// TIA Portal project "Tes simulation extract_V15.1" (V15.1)

(* hardware
DEVICE "S71500/ET200MP station_1"  S7-1500 station
   slot 0: "Rail_0"  Rack  6ES7 590-1***0-0AA0
   slot 1: "PLC_1"  CPU 1511-1 PN  6ES7 511-1AK01-0AB0  V2.1
      slot 3: "CPU display_1"  6ES7591-1AA00-0AA0
DEVICE "PC station"  SIMATIC PC station
   slot 0: "PC station"  Rail  SIMATIC PC-Station  V1.0
      slot 125: "Stationmanager"  Station_Manager  V6.0.4
   slot 1: "IE general_1"  IE General  IE_CP  V8.2.0
   slot 2: "HMI_RT_1"  WinCC RT Advanced  6AV2 104-0xxxx-xxxx  15.1.0.0
      slot 33792: "Host interface"  Host interface
*)

// ===== PLC "PLC_1"  CPU 1511-1 PN =====

VAR_GLOBAL   // PLC tag table "Default tag table"
   "Clock_Byte" AT %MB0 : Byte;
   "Clock_10Hz" AT %M0.0 : Bool;
   "Clock_5Hz" AT %M0.1 : Bool;
   "Clock_2.5Hz" AT %M0.2 : Bool;
   "Clock_2Hz" AT %M0.3 : Bool;
   "Clock_1.25Hz" AT %M0.4 : Bool;
   "Clock_1Hz" AT %M0.5 : Bool;
   "Clock_0.625Hz" AT %M0.6 : Bool;
   "Clock_0.5Hz" AT %M0.7 : Bool;
   "Start Preparation V1" AT %M100.0 : Bool;
   "Pressure Vesel" AT %MW200 : Word;
   "Pressure Steam" AT %MW230 : Int;
   "Tag_3" AT %MW1 : Word;
   "Tag_4" AT %MB1 : Byte;
   "Tag_5" AT %T1 : Timer;
   "Tag_2" AT %T2 : Timer;
   "Tag_6" AT %MB26 : Byte;
   "Tag_7" AT %T3 : Timer;
   "Tag_8" AT %T4 : Timer;
   "Tag_9" AT %T5 : Timer;
   "Tag_10" AT %M100.1 : Bool;
   "Tag_11" AT %T6 : Timer;
   "Tag_12" AT %T7 : Timer;
   "START Proses" AT %M100.2 : Bool;
   "Tag_13" AT %T8 : Timer;
   "Tag_14" AT %MB4 : Byte;
   "Tag_15" AT %T9 : Timer;
   "Tag_16" AT %MB8 : Byte;
   "Tag_17" AT %MB6 : Byte;
   "Tag_18" AT %T10 : Timer;
   "START SUPPLY" AT %M100.3 : Bool;
   "Tag_20" AT %T11 : Timer;
   "TEMP SENSOR 1" AT %MW164 : Word;
   "Tag_21" AT %T12 : Timer;
   "TEMP SENSOR 2" AT %MW166 : Int;
   "Tag_22" AT %MB30 : Byte;
   "START PROSES V1" AT %M100.4 : Bool;
   "Tag_19" AT %MW2 : Int;
   "TEMPERATURE VESSEL 1" AT %MW240 : Int;
   "Tag_23" AT %MB2 : Byte;
   "Tag_24" AT %T13 : Timer;
   "Tag_25" AT %T14 : Timer;
   "Tag_26" AT %T15 : Timer;
   "Tag_27" AT %T16 : Timer;
   "Tag_28" AT %T17 : Timer;
   "Tag_29" AT %T18 : Timer;
   "Tag_30" AT %T19 : Timer;
   "Tag_31" AT %T20 : Timer;
   "Tag_32" AT %T21 : Timer;
   "Tag_33" AT %T22 : Timer;
   "Count Preparation V1" AT %MW120 : Int;
   "Count Step Proses V1" AT %MW140 : Int;
   "START TRANSFER" AT %M100.5 : Bool;
   "Tag_36" AT %M30.4 : Bool;
   "Tag_37" AT %T23 : Timer;
   "Tag_38" AT %T24 : Timer;
   "Tag_39" AT %T35 : Timer;
   "Tag_40" AT %T25 : Timer;
   "Tag_41" AT %T26 : Timer;
   "START PROSES V2" AT %M100.6 : Bool;
   "Pressure Vessel 2" AT %MW202 : Int;
   "TEMPERATURE VESSEL 2" AT %MW242 : Int;
   "Tag_42" AT %T27 : Timer;
   "Tag_43" AT %T28 : Timer;
   "Tag_44" AT %T29 : Timer;
   "Tag_45" AT %T30 : Timer;
   "Tag_46" AT %T31 : Timer;
   "Tag_47" AT %T32 : Timer;
   "Tag_48" AT %T33 : Timer;
   "Tag_49" AT %T34 : Timer;
   "Tag_50" AT %T36 : Timer;
   "Count Step Proses V2" AT %MW142 : Int;
   "Tag_52" AT %MB5 : Byte;
   "Start Preparation V7" AT %M102.0 : Bool;
   "Tag_54" AT %M102.1 : Bool;
   "START PROSES V3" AT %M100.7 : Bool;
   "Tag_55" AT %T38 : Timer;
   "Pressure Vessel 3" AT %MW204 : Int;
   "TEMPERATURE VESSEL 3" AT %MW244 : Int;
   "Tag_56" AT %T39 : Timer;
   "Tag_57" AT %T40 : Timer;
   "Tag_58" AT %T41 : Timer;
   "Tag_59" AT %T42 : Timer;
   "Tag_60" AT %T43 : Timer;
   "Tag_61" AT %T44 : Timer;
   "Tag_62" AT %T45 : Timer;
   "Tag_63" AT %T46 : Timer;
   "Tag_64" AT %T47 : Timer;
   "Count Step Proses V3" AT %MW144 : Int;
   "Tag_66" AT %MB9 : Byte;
   "Tag_67" AT %M102.2 : Bool;
   "Start Proses V4" AT %M101.0 : Bool;
   "Pressure Vessel 4" AT %MW206 : Int;
   "Tag_69" AT %T48 : Timer;
   "TEMPERATURE VESSEL 4" AT %MW246 : Int;
   "Tag_70" AT %T49 : Timer;
   "Tag_71" AT %T50 : Timer;
   "Tag_72" AT %T51 : Timer;
   "Tag_73" AT %T52 : Timer;
   "Tag_74" AT %T53 : Timer;
   "Tag_75" AT %T54 : Timer;
   "Tag_76" AT %T55 : Timer;
   "Tag_77" AT %T56 : Timer;
   "Tag_78" AT %T57 : Timer;
   "Count Step Proses V4" AT %MW146 : Int;
   "Tag_80" AT %MB12 : Byte;
   "Tag_81" AT %MB13 : Byte;
   "Pressure vessel 5" AT %MW208 : Int;
   "TEMPERATURE VESSEL 5" AT %MW248 : Int;
   "START PROSES V5" AT %M101.1 : Bool;
   "Tag_82" AT %M102.3 : Bool;
   "Tag_83" AT %T58 : Timer;
   "Tag_84" AT %T59 : Timer;
   "Tag_85" AT %T60 : Timer;
   "Tag_86" AT %T61 : Timer;
   "Tag_87" AT %T62 : Timer;
   "Tag_88" AT %T63 : Timer;
   "Tag_89" AT %T64 : Timer;
   "Tag_90" AT %T65 : Timer;
   "Tag_91" AT %T66 : Timer;
   "Tag_92" AT %T67 : Timer;
   "Count Step Proses V5" AT %MW148 : Int;
   "Pressure Vessel 6" AT %MW210 : Int;
   "TEMPERATURE VESSEL 6" AT %MW250 : Int;
   "Tag_94" AT %T68 : Timer;
   "Tag_95" AT %M102.4 : Bool;
   "Tag_96" AT %T69 : Timer;
   "Tag_97" AT %T70 : Timer;
   "Tag_98" AT %T71 : Timer;
   "Tag_99" AT %T72 : Timer;
   "Tag_100" AT %T73 : Timer;
   "Tag_101" AT %T74 : Timer;
   "Tag_102" AT %T75 : Timer;
   "Tag_103" AT %T76 : Timer;
   "Tag_104" AT %T77 : Timer;
   "Tag_105" AT %MB20 : Byte;
   "Tag_106" AT %MB21 : Byte;
   "START PROSES V6" AT %M101.2 : Bool;
   "Pressure Vessel 7" AT %MW212 : Int;
   "TEMPERATURE VESSEL 7" AT %MW252 : Int;
   "Tag_107" AT %T78 : Timer;
   "Tag_108" AT %M102.5 : Bool;
   "Tag_109" AT %T79 : Timer;
   "Tag_110" AT %T80 : Timer;
   "Tag_111" AT %T81 : Timer;
   "Tag_112" AT %T82 : Timer;
   "Tag_113" AT %T83 : Timer;
   "Tag_114" AT %T84 : Timer;
   "Tag_115" AT %T85 : Timer;
   "Tag_116" AT %T86 : Timer;
   "Tag_117" AT %T87 : Timer;
   "Tag_118" AT %MB24 : Byte;
   "Tag_119" AT %MB25 : Byte;
   "Start preparation v2" AT %M101.3 : Bool;
   "Tag_1" AT %T88 : Timer;
   "Tag_120" AT %T90 : Timer;
   "Tag_121" AT %T91 : Timer;
   "Tag_122" AT %T92 : Timer;
   "Tag_123" AT %T93 : Timer;
   "Tag_124" AT %T94 : Timer;
   "Tag_125" AT %T95 : Timer;
   "Count Preparation V2" AT %MW122 : Int;
   "Start Preparation v3" AT %M101.4 : Bool;
   "Tag_127" AT %T96 : Timer;
   "Tag_128" AT %T97 : Timer;
   "Tag_129" AT %T98 : Timer;
   "Tag_130" AT %T99 : Timer;
   "Tag_131" AT %T100 : Timer;
   "Tag_132" AT %T101 : Timer;
   "Tag_133" AT %T102 : Timer;
   "Count Preparation V3" AT %MW124 : Int;
   "Start Preparation V4" AT %M101.5 : Bool;
   "Tag_135" AT %T103 : Timer;
   "Tag_136" AT %T104 : Timer;
   "Tag_137" AT %T105 : Timer;
   "Tag_138" AT %T106 : Timer;
   "Tag_139" AT %T107 : Timer;
   "Tag_140" AT %T108 : Timer;
   "Tag_141" AT %T109 : Timer;
   "Count Preparation V4" AT %MW126 : Int;
   "Tag_143" AT %MW1226 : Int;
   "Start Preparation V5" AT %M101.6 : Bool;
   "Tag_144" AT %T110 : Timer;
   "Tag_145" AT %T111 : Timer;
   "Tag_146" AT %T112 : Timer;
   "Tag_147" AT %T113 : Timer;
   "Tag_148" AT %T114 : Timer;
   "Tag_149" AT %T115 : Timer;
   "Tag_150" AT %T116 : Timer;
   "Tag_151" AT %MB16 : Byte;
   "Start Preparation V6" AT %M101.7 : Bool;
   "Tag_152" AT %T117 : Timer;
   "Tag_153" AT %T118 : Timer;
   "Tag_154" AT %T119 : Timer;
   "Tag_155" AT %T120 : Timer;
   "Tag_156" AT %T121 : Timer;
   "Tag_157" AT %T122 : Timer;
   "Tag_158" AT %T123 : Timer;
   "Count Preparation V5" AT %MW128 : Int;
   "Count Preparation V6" AT %MW130 : Int;
   "Tag_53" AT %M102.6 : Bool;
   "Tag_161" AT %T124 : Timer;
   "Tag_162" AT %T125 : Timer;
   "Tag_163" AT %T126 : Timer;
   "Tag_164" AT %T127 : Timer;
   "Tag_165" AT %T128 : Timer;
   "Tag_166" AT %T129 : Timer;
   "Tag_167" AT %T130 : Timer;
   "Count Preparation V7" AT %MW132 : Int;
   "Tag_169" AT %MW134 : Int;
   "Count Step Proses V6" AT %MW150 : Int;
   "Count Step Proses V7" AT %MW152 : Int;
   "Tag_35" AT %MW2244 : Int;
   "START PROSES V7" AT %M102.7 : Bool;
   "Tag_51" AT %MB17 : Byte;
   "Tag_65" AT %T131 : Timer;
   "Tag_68" AT %T132 : Timer;
   "Tag_79" AT %T133 : Timer;
   "Tag_93" AT %T134 : Timer;
   "Tag_170" AT %MW40 : Word;
   "Tag_171" AT %T135 : Timer;
   "Reset Cycle" AT %M103.0 : Bool;
   "Tag_34" AT %T136 : Timer;
   "Tag_126" AT %T137 : Timer;
   "Tag_134" AT %T138 : Timer;
   "Tag_142" AT %T139 : Timer;
   "Tag_159" AT %T140 : Timer;
   "Tag_160" AT %T141 : Timer;
   "Tag_168" AT %T142 : Timer;
   "Tag_172" AT %M1.1 : Bool;
   "Tag_173" AT %M1.0 : Bool;
   "Tag_174" AT %T143 : Timer;
   "Tag_175" AT %T144 : Timer;
   "Tag_176" AT %T145 : Timer;
   "Tag_177" AT %T146 : Timer;
   "Tag_178" AT %T147 : Timer;
   "Tag_179" AT %T148 : Timer;
   "Tag_180" AT %T149 : Timer;
   "Tag_181" AT %T150 : Timer;
   "Tag_182" AT %T151 : Timer;
   "Tag_183" AT %M4.0 : Bool;
   "Tag_184" AT %M8.0 : Bool;
   "Tag_185" AT %M12.0 : Bool;
   "Tag_186" AT %M16.0 : Bool;
   "Tag_187" AT %M20.0 : Bool;
   "Tag_188" AT %M24.0 : Bool;
   "Tag_189" AT %M30.5 : Bool;
   "Tag_190" AT %M30.7 : Bool;
   "Emergency" AT %M103.1 : Bool;
   "Tag_191" AT %MW4 : Word;
   "Tag_192" AT %MW8 : Word;
   "Tag_193" AT %MW12 : Word;
   "Tag_194" AT %MW16 : Word;
   "Tag_195" AT %MW20 : Word;
   "Tag_196" AT %MW24 : Word;
   "Tag_197" AT %MW26 : Word;
   "Tag_198" AT %MW30 : Word;
   "Tag_199" AT %MW160 : Int;
   "Tag_200" AT %MW243 : Int;
END_VAR

DATA_BLOCK "DB10"   // DB10
{ S7_Optimized_Access := 'FALSE' }
VERSION : 0.1
   VAR
      Pulse_1 : Bool;
      Pulse_2 : Bool;
      Pulse_3 : Bool;
      Pulse_4 : Bool;
      Pulse_5 : Bool;
      Pulse_6 : Bool;
      Pulse_7 : Bool;
      Pulse_8 : Bool;
      Pulse_9 : Bool;
      Pulse_10 : Bool;
      Pulse_11 : Bool;
      Pulse_12 : Bool;
      Pulse_13 : Bool;
      Pulse_14 : Bool;
      Pulse_15 : Bool;
      Pulse_16 : Bool;
      Pulse_17 : Bool;
      Pulse_18 : Bool;
      Pulse_19 : Bool;
      Pulse_20 : Bool;
      Pulse_21 : Bool;
      Pulse_22 : Bool;
      Pulse_23 : Bool;
      Pulse_24 : Bool;
      Pulse_25 : Bool;
      Pulse_26 : Bool;
      Pulse_27 : Bool;
      Pulse_28 : Bool;
      Pulse_29 : Bool;
      Pulse_30 : Bool;
      Pulse_31 : Bool;
      Pulse_32 : Bool;
      Pulse_33 : Bool;
      Pulse_34 : Bool;
      Pulse_35 : Bool;
      Pulse_36 : Bool;
      Pulse_37 : Bool;
      Pulse_38 : Bool;
      Pulse_39 : Bool;
      Pulse_40 : Bool;
      Pulse_41 : Bool;
      Pulse_42 : Bool;
      Pulse_43 : Bool;
      Pulse_44 : Bool;
      Pulse_45 : Bool;
      Pulse_46 : Bool;
      Pulse_47 : Bool;
      Pulse_48 : Bool;
      Pulse_49 : Bool;
      Pulse_50 : Bool;
      Pulse_51 : Bool;
      Pulse_52 : Bool;
      Pulse_53 : Bool;
      Pulse_54 : Bool;
      Pulse_55 : Bool;
      Pulse_56 : Bool;
      Pulse_57 : Bool;
      Pulse_58 : Bool;
      Pulse_59 : Bool;
      Pulse_60 : Bool;
      Pulse_61 : Bool;
      Pulse_62 : Bool;
      Pulse_63 : Bool;
      Pulse_64 : Bool;
      Pulse_65 : Bool;
      Pulse_66 : Bool;
      Pulse_67 : Bool;
      Pulse_68 : Bool;
      Pulse_69 : Bool;
      Pulse_70 : Bool;
      Pulse_71 : Bool;
      Pulse_72 : Bool;
      Pulse_73 : Bool;
      Pulse_74 : Bool;
      Pulse_75 : Bool;
      Pulse_76 : Bool;
      Pulse_77 : Bool;
      Pulse_78 : Bool;
      Pulse_79 : Bool;
      Pulse_80 : Bool;
      Pulse_81 : Bool;
      Pulse_82 : Bool;
      Pulse_83 : Bool;
      Pulse_84 : Bool;
      Pulse_85 : Bool;
      Pulse_86 : Bool;
      Pulse_87 : Bool;
      Pulse_88 : Bool;
      Pulse_89 : Bool;
      Pulse_90 : Bool;
      Pulse_91 : Bool;
      Pulse_92 : Bool;
      Pulse_93 : Bool;
      Pulse_94 : Bool;
      Pulse_95 : Bool;
      Pulse_96 : Bool;
      Pulse_97 : Bool;
      Pulse_98 : Bool;
      Pulse_99 : Bool;
      Pulse_100 : Bool;
      Pulse_101 : Bool;
      Pulse_102 : Bool;
      Pulse_103 : Bool;
      Pulse_104 : Bool;
      Pulse_105 : Bool;
      Pulse_106 : Bool;
      Pulse_107 : Bool;
      Pulse_108 : Bool;
      Pulse_109 : Bool;
      Pulse_110 : Bool;
      Pulse_111 : Bool;
      Pulse_112 : Bool;
      Pulse_113 : Bool;
      Pulse_114 : Bool;
      Pulse_115 : Bool;
      Pulse_116 : Bool;
      Pulse_117 : Bool;
      Pulse_118 : Bool;
      Pulse_119 : Bool;
      Pulse_120 : Bool;
      Pulse_121 : Bool;
      Pulse_122 : Bool;
      Pulse_123 : Bool;
      Pulse_124 : Bool;
      Pulse_125 : Bool;
      Pulse_126 : Bool;
      Pulse_127 : Bool;
      Pulse_128 : Bool;
      Pulse_129 : Bool;
      Pulse_130 : Bool;
      Pulse_131 : Bool;
      Pulse_132 : Bool;
      Pulse_133 : Bool;
      Pulse_134 : Bool;
      Pulse_135 : Bool;
      Pulse_136 : Bool;
      Pulse_137 : Bool;
      Pulse_138 : Bool;
      Pulse_139 : Bool;
      Pulse_140 : Bool;
      Pulse_141 : Bool;
      Pulse_142 : Bool;
      Pulse_143 : Bool;
      Pulse_144 : Bool;
      Pulse_145 : Bool;
      Pulse_146 : Bool;
      Pulse_147 : Bool;
      Pulse_148 : Bool;
      Pulse_149 : Bool;
      Pulse_150 : Bool;
      Pulse_151 : Bool;
      Pulse_152 : Bool;
      Pulse_153 : Bool;
      Pulse_154 : Bool;
      Pulse_155 : Bool;
      Pulse_156 : Bool;
      Pulse_157 : Bool;
      Pulse_158 : Bool;
      Pulse_159 : Bool;
      Pulse_160 : Bool;
      Pulse_161 : Bool;
      Pulse_162 : Bool;
      Pulse_163 : Bool;
      Pulse_164 : Bool;
      Pulse_165 : Bool;
      Pulse_166 : Bool;
      Pulse_167 : Bool;
      Pulse_168 : Bool;
      Pulse_169 : Bool;
      Pulse_170 : Bool;
      Pulse_171 : Bool;
      Pulse_172 : Bool;
      Pulse_173 : Bool;
      Pulse_174 : Bool;
      Pulse_175 : Bool;
      Pulse_176 : Bool;
      Pulse_177 : Bool;
      Pulse_178 : Bool;
      Pulse_179 : Bool;
      Pulse_180 : Bool;
      Pulse_181 : Bool;
      Pulse_182 : Bool;
      Pulse_183 : Bool;
      Pulse_184 : Bool;
      Pulse_185 : Bool;
      Pulse_186 : Bool;
      Pulse_187 : Bool;
      Pulse_188 : Bool;
      Pulse_189 : Bool;
      Pulse_190 : Bool;
      Pulse_191 : Bool;
      Pulse_192 : Bool;
      Pulse_193 : Bool;
      Pulse_194 : Bool;
      Pulse_195 : Bool;
      Pulse_196 : Bool;
      Pulse_197 : Bool;
      Pulse_198 : Bool;
      Pulse_199 : Bool;
      Pulse_200 : Bool;
      Pulse_201 : Array[0..100] of Bool;
   END_VAR
BEGIN
END_DATA_BLOCK

DATA_BLOCK "DB11"   // DB11
{ S7_Optimized_Access := 'FALSE' }
VERSION : 0.1
   VAR
      pressureSteamStatus : Bool;
      pressureVeselStatus : Bool;
      "TANK FLAVOUR" : Bool;
      "TANK HIDROLIC" : Bool;
      CycleCounter : Int;
      ReStart_V1 : Bool;
      ReStart_V2 : Bool;
      ReStart_V3 : Bool;
      ReStart_V4 : Bool;
      ReStart_V5 : Bool;
      ReStart_V6 : Bool;
      ReStart_V7 : Bool;
      Mode : Bool;
      NextVessel : Bool;
      Finish_V1 : Bool;
      Finish_V2 : Bool;
      Finish_V3 : Bool;
      Finish_V4 : Bool;
      Finish_V5 : Bool;
      Finish_V6 : Bool;
      Finish_V7 : Bool;
      Terisi_V1 : Bool;
      Terisi_V2 : Bool;
      Terisi_V3 : Bool;
      Terisi_V4 : Bool;
      Terisi_V5 : Bool;
      Terisi_V6 : Bool;
      Terisi_V7 : Bool;
      Start_VP_PumpFlavour : Bool;
      Start_VP_PumpHidrolic : Bool;
      Stop_VP_PumpFlavour : Bool;
      Sstop_VP_PumpHidrolic : Bool;
   END_VAR
BEGIN
END_DATA_BLOCK

DATA_BLOCK "DB99"   // DB99
{ S7_Optimized_Access := 'TRUE' }
VERSION : 0.1
// stored: InstanceOfName Step_Generator
"Step_Generator"
BEGIN
END_DATA_BLOCK

DATA_BLOCK "DB100"   // DB100
{ S7_Optimized_Access := 'TRUE' }
VERSION : 0.1
// stored: InstanceOfName Step_Generator
"Step_Generator"
BEGIN
END_DATA_BLOCK

DATA_BLOCK "DB101"   // DB101
{ S7_Optimized_Access := 'TRUE' }
VERSION : 0.1
// stored: InstanceOfName Step_Generator
"Step_Generator"
BEGIN
END_DATA_BLOCK

DATA_BLOCK "DB102"   // DB102
{ S7_Optimized_Access := 'TRUE' }
VERSION : 0.1
// stored: InstanceOfName Step_Generator
"Step_Generator"
BEGIN
END_DATA_BLOCK

DATA_BLOCK "DB103"   // DB103
{ S7_Optimized_Access := 'TRUE' }
VERSION : 0.1
// stored: InstanceOfName Step_Generator
"Step_Generator"
BEGIN
END_DATA_BLOCK

DATA_BLOCK "DB104"   // DB104
{ S7_Optimized_Access := 'TRUE' }
VERSION : 0.1
// stored: InstanceOfName Step_Generator
"Step_Generator"
BEGIN
END_DATA_BLOCK

DATA_BLOCK "DB105"   // DB105
{ S7_Optimized_Access := 'TRUE' }
VERSION : 0.1
// stored: InstanceOfName Step_Generator
"Step_Generator"
BEGIN
END_DATA_BLOCK

DATA_BLOCK "DB106"   // DB106
{ S7_Optimized_Access := 'TRUE' }
VERSION : 0.1
// stored: InstanceOfName Step_Generator
"Step_Generator"
BEGIN
END_DATA_BLOCK

DATA_BLOCK "DB107"   // DB107
{ S7_Optimized_Access := 'TRUE' }
VERSION : 0.1
// stored: InstanceOfName Step_Generator
"Step_Generator"
BEGIN
END_DATA_BLOCK

DATA_BLOCK "DB108"   // DB108
{ S7_Optimized_Access := 'TRUE' }
VERSION : 0.1
// stored: InstanceOfName Step_Generator
"Step_Generator"
BEGIN
END_DATA_BLOCK

DATA_BLOCK "DB109"   // DB109
{ S7_Optimized_Access := 'TRUE' }
VERSION : 0.1
// stored: InstanceOfName Step_Generator
"Step_Generator"
BEGIN
END_DATA_BLOCK

DATA_BLOCK "DB110"   // DB110
{ S7_Optimized_Access := 'TRUE' }
VERSION : 0.1
// stored: InstanceOfName Step_Generator
"Step_Generator"
BEGIN
END_DATA_BLOCK

DATA_BLOCK "DB111"   // DB111
{ S7_Optimized_Access := 'TRUE' }
VERSION : 0.1
// stored: InstanceOfName Step_Generator
"Step_Generator"
BEGIN
END_DATA_BLOCK

DATA_BLOCK "DB112"   // DB112
{ S7_Optimized_Access := 'TRUE' }
VERSION : 0.1
// stored: InstanceOfName Step_Generator
"Step_Generator"
BEGIN
END_DATA_BLOCK

DATA_BLOCK "DB113"   // DB113
{ S7_Optimized_Access := 'TRUE' }
VERSION : 0.1
// stored: InstanceOfName Step_Generator
"Step_Generator"
BEGIN
END_DATA_BLOCK

DATA_BLOCK "DB114"   // DB114
{ S7_Optimized_Access := 'TRUE' }
VERSION : 0.1
// stored: InstanceOfName Step_Generator
"Step_Generator"
BEGIN
END_DATA_BLOCK

DATA_BLOCK "DB115"   // DB115
{ S7_Optimized_Access := 'TRUE' }
VERSION : 0.1
// stored: InstanceOfName Step_Generator
"Step_Generator"
BEGIN
END_DATA_BLOCK

DATA_BLOCK "DB116"   // DB116
{ S7_Optimized_Access := 'TRUE' }
VERSION : 0.1
// stored: InstanceOfName Step_Generator
"Step_Generator"
BEGIN
END_DATA_BLOCK

FUNCTION_BLOCK "Step_Generator"   // FB100, LAD
{ S7_Optimized_Access := 'TRUE' }
VERSION : 0.1
   VAR_INPUT
      En_Step_0 : Bool;
      En_Step_1 : Bool;
      En_Step_2 : Bool;
      En_Step_3 : Bool;
      En_Step_4 : Bool;
      En_Step_5 : Bool;
      En_Step_6 : Bool;
      En_Step_7 : Bool;
      En_Step_8 : Bool;
      En_Step_9 : Bool;
      En_Step_10 : Bool;
      En_Step_11 : Bool;
      En_Step_12 : Bool;
      En_Step_13 : Bool;
      En_Step_14 : Bool;
      En_Step_15 : Bool;
      En_Step_16 : Bool;
      En_Step_17 : Bool;
      En_Step_18 : Bool;
      En_Step_19 : Bool;
      En_Step_20 : Bool;
      En_Step_21 : Bool;
      En_Step_22 : Bool;
      En_Step_23 : Bool;
      En_Step_24 : Bool;
      En_Step_25 : Bool;
      En_Step_26 : Bool;
      En_Step_27 : Bool;
      En_Step_28 : Bool;
      En_Step_29 : Bool;
      En_Step_30 : Bool;
   END_VAR
   VAR_OUTPUT
      Out_Step_0 : Bool;
      Out_Step_1 : Bool;
      Out_Step_2 : Bool;
      Out_Step_3 : Bool;
      Out_Step_4 : Bool;
      Out_Step_5 : Bool;
      Out_Step_6 : Bool;
      Out_Step_7 : Bool;
      Out_Step_8 : Bool;
      Out_Step_9 : Bool;
      Out_Step_10 : Bool;
      Out_Step_11 : Bool;
      Out_Step_12 : Bool;
      Out_Step_13 : Bool;
      Out_Step_14 : Bool;
      Out_Step_15 : Bool;
      Out_Step_16 : Bool;
      Out_Step_17 : Bool;
      Out_Step_18 : Bool;
      Out_Step_19 : Bool;
      Out_Step_20 : Bool;
      Out_Step_21 : Bool;
      Out_Step_22 : Bool;
      Out_Step_23 : Bool;
      Out_Step_24 : Bool;
      Out_Step_25 : Bool;
      Out_Step_26 : Bool;
      Out_Step_27 : Bool;
      Out_Step_28 : Bool;
      Out_Step_29 : Bool;
      Out_Step_30 : Bool;
   END_VAR
   VAR_IN_OUT
      StepCounter : Int;
   END_VAR
BEGIN

REGION Network 1 (STL): Step 0 - 9
   //      A     #En_Step_0
   //      L     0
   //      T     #StepCounter
   //      L     #StepCounter
   //      L     0
   //      ==I
   //      =     #Out_Step_0
   //
   //      A     #En_Step_1
   //      L     1
   //      T     #StepCounter
   //      L     #StepCounter
   //      L     1
   //      =     #Out_Step_1
   //
   //      A     #En_Step_2
   //      L     2
   //      T     #StepCounter
   //      L     #StepCounter
   //      L     2
   //      =     #Out_Step_2
   //      A     #En_Step_3
   //      L     3
   //      T     #StepCounter
   //      =     #Out_Step_3
   //      A     #En_Step_4
   //      L     4
   //      T     #StepCounter
   //      =     #Out_Step_4
   //      A     #En_Step_5
   //      L     5
   //      T     #StepCounter
   //      =     #Out_Step_5
   //      A     #En_Step_6
   //      L     6
   //      T     #StepCounter
   //      =     #Out_Step_6
   //      A     #En_Step_7
   //      L     7
   //      T     #StepCounter
   //      =     #Out_Step_7
   //      A     #En_Step_8
   //      L     8
   //      T     #StepCounter
   //      =     #Out_Step_8
   //      A     #En_Step_9
   //      L     9
   //      T     #StepCounter
   //      =     #Out_Step_9
   //      A     #En_Step_10
   //      L     10
   //      T     #StepCounter
   //      =     #Out_Step_10
   //      A     #En_Step_11
   //      L     11
   //      T     #StepCounter
   //      =     #Out_Step_11
   //      A     #En_Step_12
   //      L     1
   //      T     #StepCounter
   //      =     #Out_Step_12
   //
   //
   //
   //
   //
   //
   //
   //
   //
   //
   //
   //
END_REGION

REGION Network 2
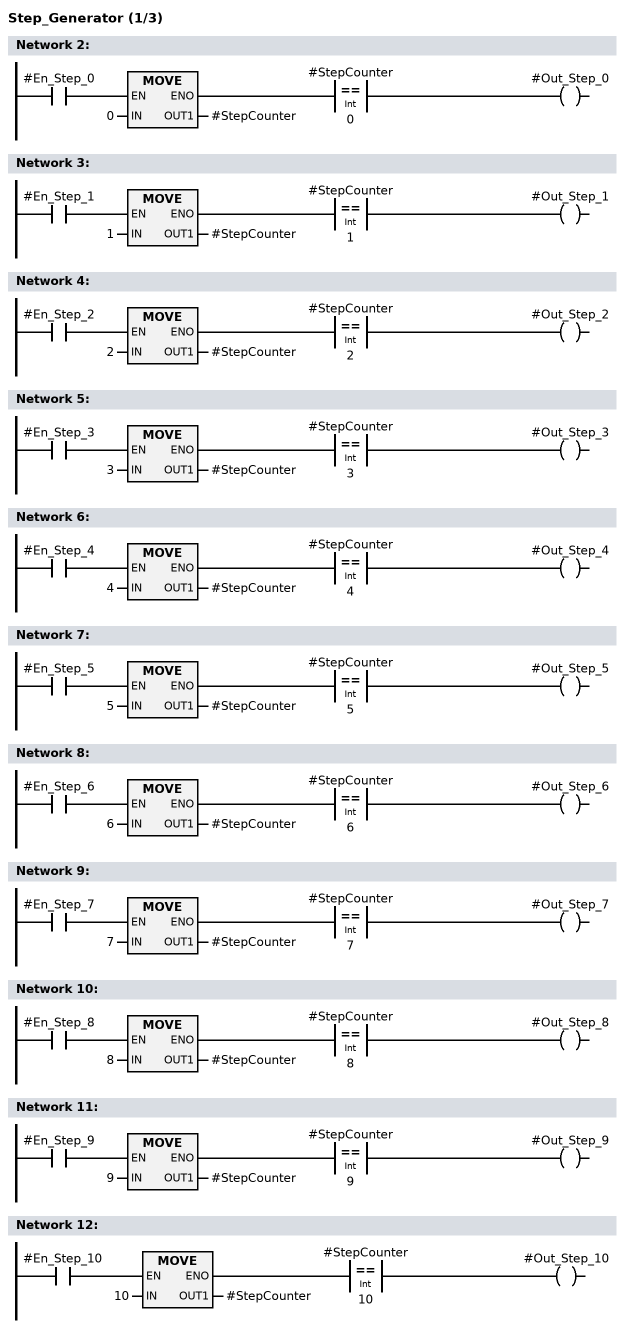
   RUNG wire#powerrail
      Contact( #En_Step_0 )
      Move(in := 0, out1 => #StepCounter)
      { S7_Templates := "SrcType := Int" } EQ_Contact(in1 := #StepCounter, in2 := 0)
      Coil( #Out_Step_0 )
   END_RUNG
   // the same network as SCL:
   IF #En_Step_0 THEN #StepCounter := 0; END_IF;
   #Out_Step_0 := #En_Step_0 AND (#StepCounter = 0);
END_REGION

REGION Network 3
   RUNG wire#powerrail
      Contact( #En_Step_1 )
      Move(in := 1, out1 => #StepCounter)
      { S7_Templates := "SrcType := Int" } EQ_Contact(in1 := #StepCounter, in2 := 1)
      Coil( #Out_Step_1 )
   END_RUNG
   // the same network as SCL:
   IF #En_Step_1 THEN #StepCounter := 1; END_IF;
   #Out_Step_1 := #En_Step_1 AND (#StepCounter = 1);
END_REGION

REGION Network 4
   RUNG wire#powerrail
      Contact( #En_Step_2 )
      Move(in := 2, out1 => #StepCounter)
      { S7_Templates := "SrcType := Int" } EQ_Contact(in1 := #StepCounter, in2 := 2)
      Coil( #Out_Step_2 )
   END_RUNG
   // the same network as SCL:
   IF #En_Step_2 THEN #StepCounter := 2; END_IF;
   #Out_Step_2 := #En_Step_2 AND (#StepCounter = 2);
END_REGION

REGION Network 5
   RUNG wire#powerrail
      Contact( #En_Step_3 )
      Move(in := 3, out1 => #StepCounter)
      { S7_Templates := "SrcType := Int" } EQ_Contact(in1 := #StepCounter, in2 := 3)
      Coil( #Out_Step_3 )
   END_RUNG
   // the same network as SCL:
   IF #En_Step_3 THEN #StepCounter := 3; END_IF;
   #Out_Step_3 := #En_Step_3 AND (#StepCounter = 3);
END_REGION

REGION Network 6
   RUNG wire#powerrail
      Contact( #En_Step_4 )
      Move(in := 4, out1 => #StepCounter)
      { S7_Templates := "SrcType := Int" } EQ_Contact(in1 := #StepCounter, in2 := 4)
      Coil( #Out_Step_4 )
   END_RUNG
   // the same network as SCL:
   IF #En_Step_4 THEN #StepCounter := 4; END_IF;
   #Out_Step_4 := #En_Step_4 AND (#StepCounter = 4);
END_REGION

REGION Network 7
   RUNG wire#powerrail
      Contact( #En_Step_5 )
      Move(in := 5, out1 => #StepCounter)
      { S7_Templates := "SrcType := Int" } EQ_Contact(in1 := #StepCounter, in2 := 5)
      Coil( #Out_Step_5 )
   END_RUNG
   // the same network as SCL:
   IF #En_Step_5 THEN #StepCounter := 5; END_IF;
   #Out_Step_5 := #En_Step_5 AND (#StepCounter = 5);
END_REGION

REGION Network 8
   RUNG wire#powerrail
      Contact( #En_Step_6 )
      Move(in := 6, out1 => #StepCounter)
      { S7_Templates := "SrcType := Int" } EQ_Contact(in1 := #StepCounter, in2 := 6)
      Coil( #Out_Step_6 )
   END_RUNG
   // the same network as SCL:
   IF #En_Step_6 THEN #StepCounter := 6; END_IF;
   #Out_Step_6 := #En_Step_6 AND (#StepCounter = 6);
END_REGION

REGION Network 9
   RUNG wire#powerrail
      Contact( #En_Step_7 )
      Move(in := 7, out1 => #StepCounter)
      { S7_Templates := "SrcType := Int" } EQ_Contact(in1 := #StepCounter, in2 := 7)
      Coil( #Out_Step_7 )
   END_RUNG
   // the same network as SCL:
   IF #En_Step_7 THEN #StepCounter := 7; END_IF;
   #Out_Step_7 := #En_Step_7 AND (#StepCounter = 7);
END_REGION

REGION Network 10
   RUNG wire#powerrail
      Contact( #En_Step_8 )
      Move(in := 8, out1 => #StepCounter)
      { S7_Templates := "SrcType := Int" } EQ_Contact(in1 := #StepCounter, in2 := 8)
      Coil( #Out_Step_8 )
   END_RUNG
   // the same network as SCL:
   IF #En_Step_8 THEN #StepCounter := 8; END_IF;
   #Out_Step_8 := #En_Step_8 AND (#StepCounter = 8);
END_REGION

REGION Network 11
   RUNG wire#powerrail
      Contact( #En_Step_9 )
      Move(in := 9, out1 => #StepCounter)
      { S7_Templates := "SrcType := Int" } EQ_Contact(in1 := #StepCounter, in2 := 9)
      Coil( #Out_Step_9 )
   END_RUNG
   // the same network as SCL:
   IF #En_Step_9 THEN #StepCounter := 9; END_IF;
   #Out_Step_9 := #En_Step_9 AND (#StepCounter = 9);
END_REGION

REGION Network 12
   RUNG wire#powerrail
      Contact( #En_Step_10 )
      Move(in := 10, out1 => #StepCounter)
      { S7_Templates := "SrcType := Int" } EQ_Contact(in1 := #StepCounter, in2 := 10)
      Coil( #Out_Step_10 )
   END_RUNG
   // the same network as SCL:
   IF #En_Step_10 THEN #StepCounter := 10; END_IF;
   #Out_Step_10 := #En_Step_10 AND (#StepCounter = 10);
END_REGION

REGION Network 13
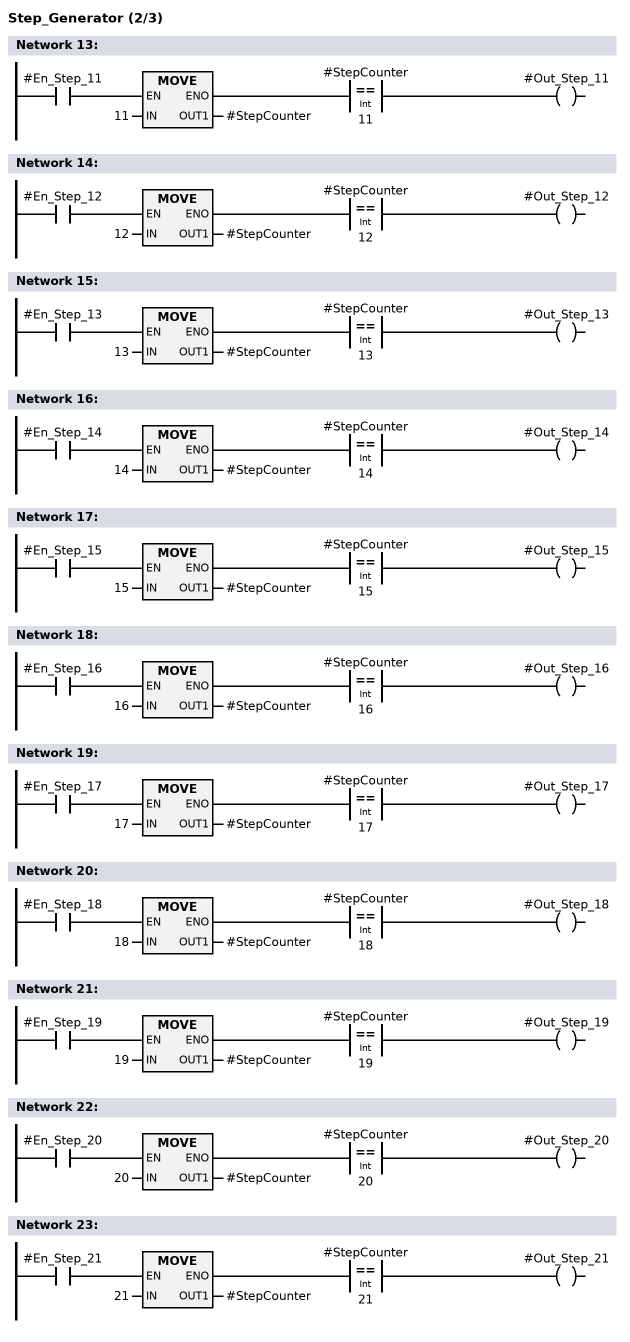
   RUNG wire#powerrail
      Contact( #En_Step_11 )
      Move(in := 11, out1 => #StepCounter)
      { S7_Templates := "SrcType := Int" } EQ_Contact(in1 := #StepCounter, in2 := 11)
      Coil( #Out_Step_11 )
   END_RUNG
   // the same network as SCL:
   IF #En_Step_11 THEN #StepCounter := 11; END_IF;
   #Out_Step_11 := #En_Step_11 AND (#StepCounter = 11);
END_REGION

REGION Network 14
   RUNG wire#powerrail
      Contact( #En_Step_12 )
      Move(in := 12, out1 => #StepCounter)
      { S7_Templates := "SrcType := Int" } EQ_Contact(in1 := #StepCounter, in2 := 12)
      Coil( #Out_Step_12 )
   END_RUNG
   // the same network as SCL:
   IF #En_Step_12 THEN #StepCounter := 12; END_IF;
   #Out_Step_12 := #En_Step_12 AND (#StepCounter = 12);
END_REGION

REGION Network 15
   RUNG wire#powerrail
      Contact( #En_Step_13 )
      Move(in := 13, out1 => #StepCounter)
      { S7_Templates := "SrcType := Int" } EQ_Contact(in1 := #StepCounter, in2 := 13)
      Coil( #Out_Step_13 )
   END_RUNG
   // the same network as SCL:
   IF #En_Step_13 THEN #StepCounter := 13; END_IF;
   #Out_Step_13 := #En_Step_13 AND (#StepCounter = 13);
END_REGION

REGION Network 16
   RUNG wire#powerrail
      Contact( #En_Step_14 )
      Move(in := 14, out1 => #StepCounter)
      { S7_Templates := "SrcType := Int" } EQ_Contact(in1 := #StepCounter, in2 := 14)
      Coil( #Out_Step_14 )
   END_RUNG
   // the same network as SCL:
   IF #En_Step_14 THEN #StepCounter := 14; END_IF;
   #Out_Step_14 := #En_Step_14 AND (#StepCounter = 14);
END_REGION

REGION Network 17
   RUNG wire#powerrail
      Contact( #En_Step_15 )
      Move(in := 15, out1 => #StepCounter)
      { S7_Templates := "SrcType := Int" } EQ_Contact(in1 := #StepCounter, in2 := 15)
      Coil( #Out_Step_15 )
   END_RUNG
   // the same network as SCL:
   IF #En_Step_15 THEN #StepCounter := 15; END_IF;
   #Out_Step_15 := #En_Step_15 AND (#StepCounter = 15);
END_REGION

REGION Network 18
   RUNG wire#powerrail
      Contact( #En_Step_16 )
      Move(in := 16, out1 => #StepCounter)
      { S7_Templates := "SrcType := Int" } EQ_Contact(in1 := #StepCounter, in2 := 16)
      Coil( #Out_Step_16 )
   END_RUNG
   // the same network as SCL:
   IF #En_Step_16 THEN #StepCounter := 16; END_IF;
   #Out_Step_16 := #En_Step_16 AND (#StepCounter = 16);
END_REGION

REGION Network 19
   RUNG wire#powerrail
      Contact( #En_Step_17 )
      Move(in := 17, out1 => #StepCounter)
      { S7_Templates := "SrcType := Int" } EQ_Contact(in1 := #StepCounter, in2 := 17)
      Coil( #Out_Step_17 )
   END_RUNG
   // the same network as SCL:
   IF #En_Step_17 THEN #StepCounter := 17; END_IF;
   #Out_Step_17 := #En_Step_17 AND (#StepCounter = 17);
END_REGION

REGION Network 20
   RUNG wire#powerrail
      Contact( #En_Step_18 )
      Move(in := 18, out1 => #StepCounter)
      { S7_Templates := "SrcType := Int" } EQ_Contact(in1 := #StepCounter, in2 := 18)
      Coil( #Out_Step_18 )
   END_RUNG
   // the same network as SCL:
   IF #En_Step_18 THEN #StepCounter := 18; END_IF;
   #Out_Step_18 := #En_Step_18 AND (#StepCounter = 18);
END_REGION

REGION Network 21
   RUNG wire#powerrail
      Contact( #En_Step_19 )
      Move(in := 19, out1 => #StepCounter)
      { S7_Templates := "SrcType := Int" } EQ_Contact(in1 := #StepCounter, in2 := 19)
      Coil( #Out_Step_19 )
   END_RUNG
   // the same network as SCL:
   IF #En_Step_19 THEN #StepCounter := 19; END_IF;
   #Out_Step_19 := #En_Step_19 AND (#StepCounter = 19);
END_REGION

REGION Network 22
   RUNG wire#powerrail
      Contact( #En_Step_20 )
      Move(in := 20, out1 => #StepCounter)
      { S7_Templates := "SrcType := Int" } EQ_Contact(in1 := #StepCounter, in2 := 20)
      Coil( #Out_Step_20 )
   END_RUNG
   // the same network as SCL:
   IF #En_Step_20 THEN #StepCounter := 20; END_IF;
   #Out_Step_20 := #En_Step_20 AND (#StepCounter = 20);
END_REGION

REGION Network 23
   RUNG wire#powerrail
      Contact( #En_Step_21 )
      Move(in := 21, out1 => #StepCounter)
      { S7_Templates := "SrcType := Int" } EQ_Contact(in1 := #StepCounter, in2 := 21)
      Coil( #Out_Step_21 )
   END_RUNG
   // the same network as SCL:
   IF #En_Step_21 THEN #StepCounter := 21; END_IF;
   #Out_Step_21 := #En_Step_21 AND (#StepCounter = 21);
END_REGION

REGION Network 24
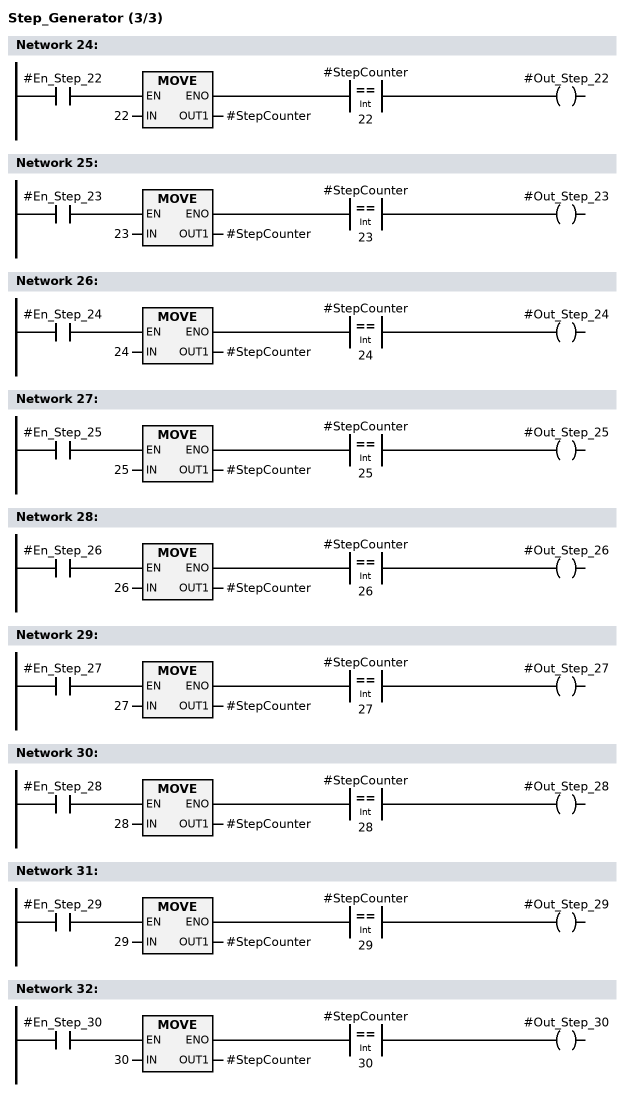
   RUNG wire#powerrail
      Contact( #En_Step_22 )
      Move(in := 22, out1 => #StepCounter)
      { S7_Templates := "SrcType := Int" } EQ_Contact(in1 := #StepCounter, in2 := 22)
      Coil( #Out_Step_22 )
   END_RUNG
   // the same network as SCL:
   IF #En_Step_22 THEN #StepCounter := 22; END_IF;
   #Out_Step_22 := #En_Step_22 AND (#StepCounter = 22);
END_REGION

REGION Network 25
   RUNG wire#powerrail
      Contact( #En_Step_23 )
      Move(in := 23, out1 => #StepCounter)
      { S7_Templates := "SrcType := Int" } EQ_Contact(in1 := #StepCounter, in2 := 23)
      Coil( #Out_Step_23 )
   END_RUNG
   // the same network as SCL:
   IF #En_Step_23 THEN #StepCounter := 23; END_IF;
   #Out_Step_23 := #En_Step_23 AND (#StepCounter = 23);
END_REGION

REGION Network 26
   RUNG wire#powerrail
      Contact( #En_Step_24 )
      Move(in := 24, out1 => #StepCounter)
      { S7_Templates := "SrcType := Int" } EQ_Contact(in1 := #StepCounter, in2 := 24)
      Coil( #Out_Step_24 )
   END_RUNG
   // the same network as SCL:
   IF #En_Step_24 THEN #StepCounter := 24; END_IF;
   #Out_Step_24 := #En_Step_24 AND (#StepCounter = 24);
END_REGION

REGION Network 27
   RUNG wire#powerrail
      Contact( #En_Step_25 )
      Move(in := 25, out1 => #StepCounter)
      { S7_Templates := "SrcType := Int" } EQ_Contact(in1 := #StepCounter, in2 := 25)
      Coil( #Out_Step_25 )
   END_RUNG
   // the same network as SCL:
   IF #En_Step_25 THEN #StepCounter := 25; END_IF;
   #Out_Step_25 := #En_Step_25 AND (#StepCounter = 25);
END_REGION

REGION Network 28
   RUNG wire#powerrail
      Contact( #En_Step_26 )
      Move(in := 26, out1 => #StepCounter)
      { S7_Templates := "SrcType := Int" } EQ_Contact(in1 := #StepCounter, in2 := 26)
      Coil( #Out_Step_26 )
   END_RUNG
   // the same network as SCL:
   IF #En_Step_26 THEN #StepCounter := 26; END_IF;
   #Out_Step_26 := #En_Step_26 AND (#StepCounter = 26);
END_REGION

REGION Network 29
   RUNG wire#powerrail
      Contact( #En_Step_27 )
      Move(in := 27, out1 => #StepCounter)
      { S7_Templates := "SrcType := Int" } EQ_Contact(in1 := #StepCounter, in2 := 27)
      Coil( #Out_Step_27 )
   END_RUNG
   // the same network as SCL:
   IF #En_Step_27 THEN #StepCounter := 27; END_IF;
   #Out_Step_27 := #En_Step_27 AND (#StepCounter = 27);
END_REGION

REGION Network 30
   RUNG wire#powerrail
      Contact( #En_Step_28 )
      Move(in := 28, out1 => #StepCounter)
      { S7_Templates := "SrcType := Int" } EQ_Contact(in1 := #StepCounter, in2 := 28)
      Coil( #Out_Step_28 )
   END_RUNG
   // the same network as SCL:
   IF #En_Step_28 THEN #StepCounter := 28; END_IF;
   #Out_Step_28 := #En_Step_28 AND (#StepCounter = 28);
END_REGION

REGION Network 31
   RUNG wire#powerrail
      Contact( #En_Step_29 )
      Move(in := 29, out1 => #StepCounter)
      { S7_Templates := "SrcType := Int" } EQ_Contact(in1 := #StepCounter, in2 := 29)
      Coil( #Out_Step_29 )
   END_RUNG
   // the same network as SCL:
   IF #En_Step_29 THEN #StepCounter := 29; END_IF;
   #Out_Step_29 := #En_Step_29 AND (#StepCounter = 29);
END_REGION

REGION Network 32
   RUNG wire#powerrail
      Contact( #En_Step_30 )
      Move(in := 30, out1 => #StepCounter)
      { S7_Templates := "SrcType := Int" } EQ_Contact(in1 := #StepCounter, in2 := 30)
      Coil( #Out_Step_30 )
   END_RUNG
   // the same network as SCL:
   IF #En_Step_30 THEN #StepCounter := 30; END_IF;
   #Out_Step_30 := #En_Step_30 AND (#StepCounter = 30);
END_REGION
END_FUNCTION_BLOCK

FUNCTION "SEQUENCE V1 PREPARATION" : Void   // FC1, LAD
{ S7_Optimized_Access := 'TRUE' }
VERSION : 0.1
   VAR_TEMP   // added for the SCL form of the ladder/FBD networks
      _w1 : Bool;
      _s5time1 : S5Time;
      _w2 : Bool;
      _s5time2 : S5Time;
   END_VAR
BEGIN

REGION Network 1: Start Preparation
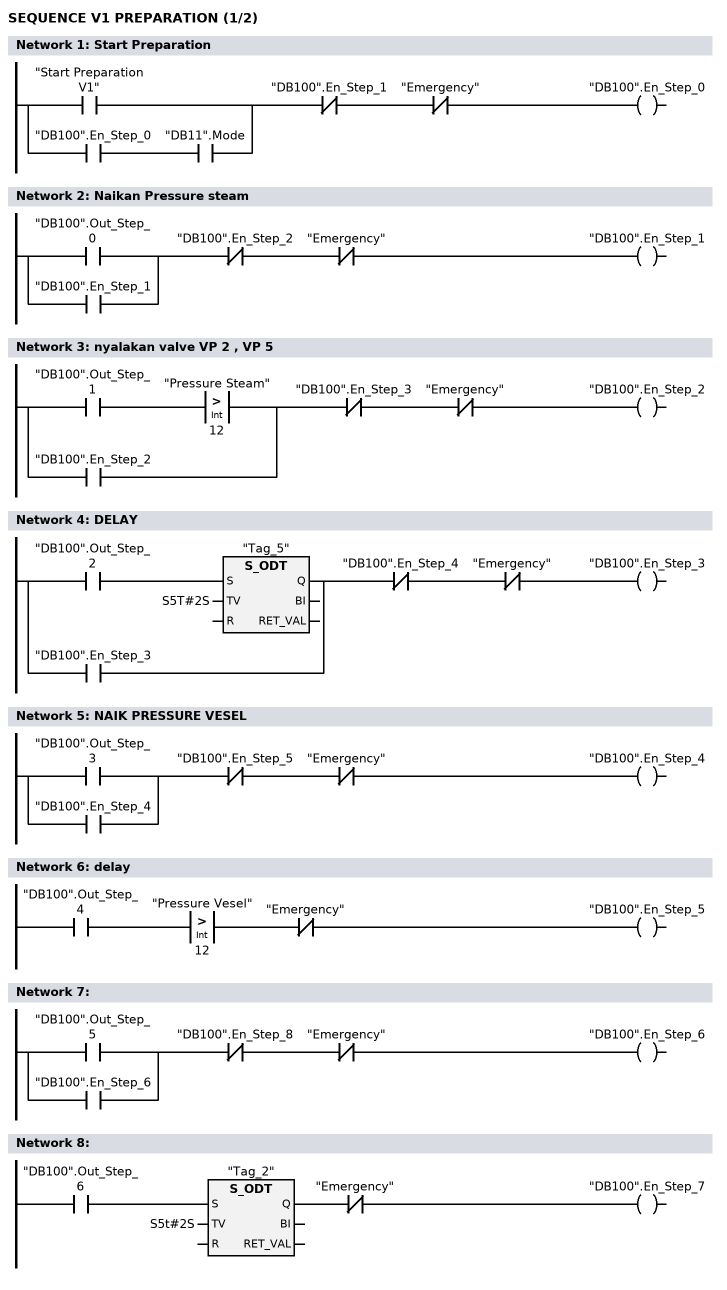
   RUNG wire#powerrail
      Contact( "Start Preparation V1" )
      wire#w1
      I_Contact( "DB100".En_Step_1 )
      I_Contact( "Emergency" )
      Coil( "DB100".En_Step_0 )
   END_RUNG
   RUNG wire#powerrail
      Contact( "DB100".En_Step_0 )
      Contact( "DB11".Mode )
   END_RUNG wire#w1
   // the same network as SCL:
   "DB100".En_Step_0 := ("Start Preparation V1" OR ("DB100".En_Step_0 AND "DB11".Mode)) AND NOT "DB100".En_Step_1 AND NOT "Emergency";
END_REGION

REGION Network 2: Naikan Pressure steam
   RUNG wire#powerrail
      Contact( "DB100".Out_Step_0 )
      wire#w1
      I_Contact( "DB100".En_Step_2 )
      I_Contact( "Emergency" )
      Coil( "DB100".En_Step_1 )
   END_RUNG
   RUNG wire#powerrail
      Contact( "DB100".En_Step_1 )
   END_RUNG wire#w1
   // the same network as SCL:
   "DB100".En_Step_1 := ("DB100".Out_Step_0 OR "DB100".En_Step_1) AND NOT "DB100".En_Step_2 AND NOT "Emergency";
END_REGION

REGION Network 3: nyalakan valve VP 2 , VP 5
   RUNG wire#powerrail
      Contact( "DB100".Out_Step_1 )
      { S7_Templates := "SrcType := Int" } GT_Contact(in1 := "Pressure Steam", in2 := 12)
      wire#w1
      I_Contact( "DB100".En_Step_3 )
      I_Contact( "Emergency" )
      Coil( "DB100".En_Step_2 )
   END_RUNG
   RUNG wire#powerrail
      Contact( "DB100".En_Step_2 )
   END_RUNG wire#w1
   // the same network as SCL:
   "DB100".En_Step_2 := (("DB100".Out_Step_1 AND ("Pressure Steam" > 12)) OR "DB100".En_Step_2) AND NOT "DB100".En_Step_3 AND NOT "Emergency";
END_REGION

REGION Network 4: DELAY
   RUNG wire#powerrail
      Contact( "DB100".Out_Step_2 )
      S_ODT(T_NO := "Tag_5", TV := S5T#2S, R :=, BI =>, RET_VAL =>)
      wire#w1
      I_Contact( "DB100".En_Step_4 )
      I_Contact( "Emergency" )
      Coil( "DB100".En_Step_3 )
   END_RUNG
   RUNG wire#powerrail
      Contact( "DB100".En_Step_3 )
   END_RUNG wire#w1
   // the same network as SCL:
   #_s5time1 := S_ODT(T_NO := "Tag_5", S := "DB100".Out_Step_2, TV := S5T#2S, Q => #_w1);
   "DB100".En_Step_3 := (#_w1 OR "DB100".En_Step_3) AND NOT "DB100".En_Step_4 AND NOT "Emergency";
END_REGION

REGION Network 5: NAIK PRESSURE VESEL
   RUNG wire#powerrail
      Contact( "DB100".Out_Step_3 )
      wire#w1
      I_Contact( "DB100".En_Step_5 )
      I_Contact( "Emergency" )
      Coil( "DB100".En_Step_4 )
   END_RUNG
   RUNG wire#powerrail
      Contact( "DB100".En_Step_4 )
   END_RUNG wire#w1
   // the same network as SCL:
   "DB100".En_Step_4 := ("DB100".Out_Step_3 OR "DB100".En_Step_4) AND NOT "DB100".En_Step_5 AND NOT "Emergency";
END_REGION

REGION Network 6: delay
   RUNG wire#powerrail
      Contact( "DB100".Out_Step_4 )
      { S7_Templates := "SrcType := Int" } GT_Contact(in1 := "Pressure Vesel", in2 := 12)
      I_Contact( "Emergency" )
      Coil( "DB100".En_Step_5 )
   END_RUNG
   // the same network as SCL:
   "DB100".En_Step_5 := "DB100".Out_Step_4 AND ("Pressure Vesel" > 12) AND NOT "Emergency";
END_REGION

REGION Network 7
   RUNG wire#powerrail
      Contact( "DB100".Out_Step_5 )
      wire#w1
      I_Contact( "DB100".En_Step_8 )
      I_Contact( "Emergency" )
      Coil( "DB100".En_Step_6 )
   END_RUNG
   RUNG wire#powerrail
      Contact( "DB100".En_Step_6 )
   END_RUNG wire#w1
   // the same network as SCL:
   "DB100".En_Step_6 := ("DB100".Out_Step_5 OR "DB100".En_Step_6) AND NOT "DB100".En_Step_8 AND NOT "Emergency";
END_REGION

REGION Network 8
   RUNG wire#powerrail
      Contact( "DB100".Out_Step_6 )
      S_ODT(T_NO := "Tag_2", TV := S5t#2S, R :=, BI =>, RET_VAL =>)
      I_Contact( "Emergency" )
      Coil( "DB100".En_Step_7 )
   END_RUNG
   // the same network as SCL:
   #_s5time1 := S_ODT(T_NO := "Tag_2", S := "DB100".Out_Step_6, TV := S5t#2S, Q => #_w1);
   "DB100".En_Step_7 := #_w1 AND NOT "Emergency";
END_REGION

REGION Network 9: TURUNKAN PRESSURE